REGION Network 21
   RUNG wire#powerrail
      { S7_Templates := "SrcType := String" } EQ_Contact(in1 := #String2, in2 := '6')
      Move(in := 125, out1 => #Decimal2_Out)
   END_RUNG
   // the same network as SCL:
   IF #String2 = '6' THEN #Decimal2_Out := 125; END_IF;
END_REGION

REGION Network 22
   RUNG wire#powerrail
      { S7_Templates := "SrcType := String" } EQ_Contact(in1 := #String2, in2 := '7')
      Move(in := 7, out1 => #Decimal2_Out)
   END_RUNG
   // the same network as SCL:
   IF #String2 = '7' THEN #Decimal2_Out := 7; END_IF;
END_REGION

REGION Network 23
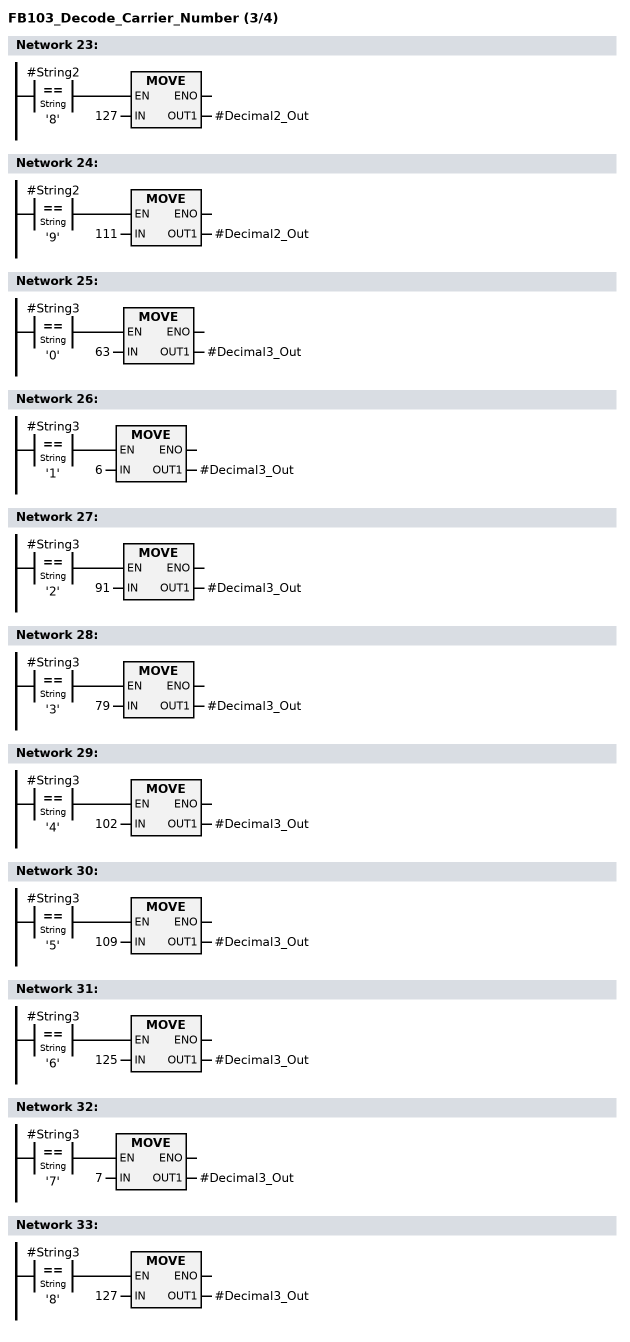
   RUNG wire#powerrail
      { S7_Templates := "SrcType := String" } EQ_Contact(in1 := #String2, in2 := '8')
      Move(in := 127, out1 => #Decimal2_Out)
   END_RUNG
   // the same network as SCL:
   IF #String2 = '8' THEN #Decimal2_Out := 127; END_IF;
END_REGION

REGION Network 24
   RUNG wire#powerrail
      { S7_Templates := "SrcType := String" } EQ_Contact(in1 := #String2, in2 := '9')
      Move(in := 111, out1 => #Decimal2_Out)
   END_RUNG
   // the same network as SCL:
   IF #String2 = '9' THEN #Decimal2_Out := 111; END_IF;
END_REGION

REGION Network 25
   RUNG wire#powerrail
      { S7_Templates := "SrcType := String" } EQ_Contact(in1 := #String3, in2 := '0')
      Move(in := 63, out1 => #Decimal3_Out)
   END_RUNG
   // the same network as SCL:
   IF #String3 = '0' THEN #Decimal3_Out := 63; END_IF;
END_REGION

REGION Network 26
   RUNG wire#powerrail
      { S7_Templates := "SrcType := String" } EQ_Contact(in1 := #String3, in2 := '1')
      Move(in := 6, out1 => #Decimal3_Out)
   END_RUNG
   // the same network as SCL:
   IF #String3 = '1' THEN #Decimal3_Out := 6; END_IF;
END_REGION

REGION Network 27
   RUNG wire#powerrail
      { S7_Templates := "SrcType := String" } EQ_Contact(in1 := #String3, in2 := '2')
      Move(in := 91, out1 => #Decimal3_Out)
   END_RUNG
   // the same network as SCL:
   IF #String3 = '2' THEN #Decimal3_Out := 91; END_IF;
END_REGION

REGION Network 28
   RUNG wire#powerrail
      { S7_Templates := "SrcType := String" } EQ_Contact(in1 := #String3, in2 := '3')
      Move(in := 79, out1 => #Decimal3_Out)
   END_RUNG
   // the same network as SCL:
   IF #String3 = '3' THEN #Decimal3_Out := 79; END_IF;
END_REGION

REGION Network 29
   RUNG wire#powerrail
      { S7_Templates := "SrcType := String" } EQ_Contact(in1 := #String3, in2 := '4')
      Move(in := 102, out1 => #Decimal3_Out)
   END_RUNG
   // the same network as SCL:
   IF #String3 = '4' THEN #Decimal3_Out := 102; END_IF;
END_REGION

REGION Network 30
   RUNG wire#powerrail
      { S7_Templates := "SrcType := String" } EQ_Contact(in1 := #String3, in2 := '5')
      Move(in := 109, out1 => #Decimal3_Out)
   END_RUNG
   // the same network as SCL:
   IF #String3 = '5' THEN #Decimal3_Out := 109; END_IF;
END_REGION

REGION Network 31
   RUNG wire#powerrail
      { S7_Templates := "SrcType := String" } EQ_Contact(in1 := #String3, in2 := '6')
      Move(in := 125, out1 => #Decimal3_Out)
   END_RUNG
   // the same network as SCL:
   IF #String3 = '6' THEN #Decimal3_Out := 125; END_IF;
END_REGION

REGION Network 32
   RUNG wire#powerrail
      { S7_Templates := "SrcType := String" } EQ_Contact(in1 := #String3, in2 := '7')
      Move(in := 7, out1 => #Decimal3_Out)
   END_RUNG
   // the same network as SCL:
   IF #String3 = '7' THEN #Decimal3_Out := 7; END_IF;
END_REGION

REGION Network 33
   RUNG wire#powerrail
      { S7_Templates := "SrcType := String" } EQ_Contact(in1 := #String3, in2 := '8')
      Move(in := 127, out1 => #Decimal3_Out)
   END_RUNG
   // the same network as SCL:
   IF #String3 = '8' THEN #Decimal3_Out := 127; END_IF;
END_REGION

REGION Network 34
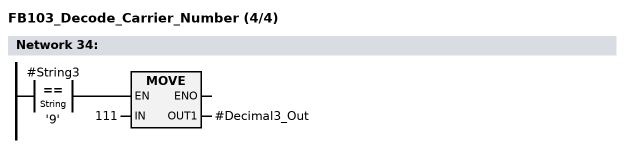
   RUNG wire#powerrail
      { S7_Templates := "SrcType := String" } EQ_Contact(in1 := #String3, in2 := '9')
      Move(in := 111, out1 => #Decimal3_Out)
   END_RUNG
   // the same network as SCL:
   IF #String3 = '9' THEN #Decimal3_Out := 111; END_IF;
END_REGION
END_FUNCTION_BLOCK

FUNCTION_BLOCK "FB104_CarrierBreakerStatus"   // FB104, LAD
{ S7_Optimized_Access := 'TRUE' }
AUTHOR : Siemens
VERSION : 1.0
// © 2018 Siemens AG 
// SIMOVE Carrier Control
   VAR
      instSystemBreakerStatus : "FB1001_EMS_BreakerStatus";
      instSystemDiagProfinet : "FB1003_LSimoveC_DiagProfinet";
      statCommunication : Bool;
      LSimoveC_DiagBreaker_Instance : "FB1001_EMS_BreakerStatus";
      LSimoveC_BreakerStatus_Instance : "FB1001_EMS_BreakerStatus";
   END_VAR
   VAR_TEMP
      tempBool_Tcc_2018_NotUsed : Bool;
   END_VAR
   VAR CONSTANT
      TCC2018_NotUsed : Bool;
   END_VAR
   VAR_TEMP   // added for the SCL form of the ladder/FBD networks
      _w1 : Bool;
   END_VAR
BEGIN

REGION Network 1: 10 System Monitoring Fuse
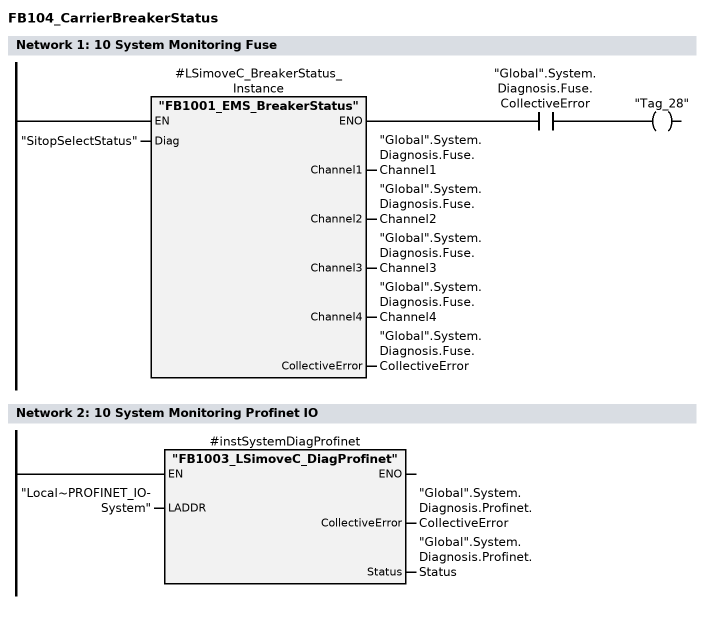
   RUNG wire#powerrail
      #LSimoveC_BreakerStatus_Instance(Diag := "SitopSelectStatus", Channel1 => "Global".System.Diagnosis.Fuse.Channel1, Channel2 => "Global".System.Diagnosis.Fuse.Channel2, Channel3 => "Global".System.Diagnosis.Fuse.Channel3, Channel4 => "Global".System.Diagnosis.Fuse.Channel4, CollectiveError => "Global".System.Diagnosis.Fuse.CollectiveError)
      Contact( "Global".System.Diagnosis.Fuse.CollectiveError )
      Coil( "Tag_28" )
   END_RUNG
   // the same network as SCL:
   #LSimoveC_BreakerStatus_Instance(Diag := "SitopSelectStatus",   // "FB1001_EMS_BreakerStatus"
                           Channel1 => "Global".System.Diagnosis.Fuse.Channel1,
                           Channel2 => "Global".System.Diagnosis.Fuse.Channel2,
                           Channel3 => "Global".System.Diagnosis.Fuse.Channel3,
                           Channel4 => "Global".System.Diagnosis.Fuse.Channel4,
                           CollectiveError => "Global".System.Diagnosis.Fuse.CollectiveError,
                           ENO => #_w1);
   "Tag_28" := #_w1 AND "Global".System.Diagnosis.Fuse.CollectiveError;
END_REGION

REGION Network 2: 10 System Monitoring Profinet IO
   RUNG wire#powerrail
      #instSystemDiagProfinet(LADDR := "Local~PROFINET_IO-System", CollectiveError => "Global".System.Diagnosis.Profinet.CollectiveError, Status => "Global".System.Diagnosis.Profinet.Status)
   END_RUNG
   // the same network as SCL:
   #instSystemDiagProfinet(LADDR := "Local~PROFINET_IO-System",   // "FB1003_LSimoveC_DiagProfinet"
                           CollectiveError => "Global".System.Diagnosis.Profinet.CollectiveError,
                           Status => "Global".System.Diagnosis.Profinet.Status);
END_REGION

REGION Network 3: 15 Navigation Transponder Antenna Left
END_REGION

REGION Network 4: 15 Navigation Transponder Antenna Right
END_REGION

REGION Network 5: 15 Navigation Identification Point
END_REGION
END_FUNCTION_BLOCK

FUNCTION_BLOCK "FB105_G120D_CarrierDrive"   // FB105, LAD
TITLE = Funkionblock for controlling a G120D
{ S7_Optimized_Access := 'FALSE' }
VERSION : 0.1
// -  ALLGEMEIN
//  - EINGÄNGE PEW
//  - STEUERWORT / CONTROLWORD
//  - ZUSTANDSWORT / STATUSWORD
//  - AUSGÄNGE PAW
//  - STÖRUNGEN
//  - ENDE
// 
// ________________________________________________________________________________
// 
// Groiß Andreas
// Siemens AG Österreich 
// Linz Kraußstraße 1-7 
// RC-AT I-IA AS-FA-SA-AE2
// 29.05.2013
// - GENERALLY
//  - INPUTS PEW
//  - STEUERWORT / CONTROLWORD
//  - ZUSTANDSWORT / STATUSWORD
//  - OUTPUTS PAW
//  - FAULTS
//  - END
// 
// ________________________________________________________________________________
// 
// Groiß Andreas
// Siemens AG Österreich 
// Linz Kraußstraße 1-7 
// I IA AS SO AP2 Surface Technology & Assembly
// 29.05.2013
   VAR_INPUT
      iPEW_ZSW1 : Word;   // IN: G120 D Zustandswort 1 / Stausword 1 PEW
      iPEW_SPEED : Word;   // IN: G120 D Aktual-Drehzahl / Actual-Speed of rotation PEW
      iPEW_INPUTS : Word;   // IN: G120 D digitale Eingänge / digital Inputs PEW
      iPEW_ERROR : Word;   // IN: G120 D Störcode / Errorcode PEW
      iEN_ERROR : Bool;   // IN: Freigabe Störmeldungen / IN: Enable Errormessages
      iON : Bool;   // IN: STW1_Bit_0 Steuerung Ein / IN: STW1_Bit_0 Control ON
      iPOWER_ON : Bool;   // IN: Kraftschalter ist EIN / IN: Power is switched on
      iENABLE : Bool;   // IN: Freigabe / IN: Enable
      iREVERSE : Bool;   // IN: STW1_Bit_11
      iBREAK : Bool;   // IN: Löse Bremse / IN: Release Break
      iDDS : Bool;   // IN: FU Datenset (0 = DDS0 / 1 = DDS1)
      iDO0 : Bool;   // IN: 1=Digitaler Ausgang aktiv/ 0=Digitaler Ausgang nicht aktiv
      iDO1 : Bool;   // IN: 1=Digitaler Ausgang aktiv/ 0=Digitaler Ausgang nicht aktiv
      iER_RESET : Bool;   // IN: Störung quittieren / IN: Error Reset
      iSET_SPEED : DInt;   // IN: Sollgeschwindigkeit in mm/min / IN: Setpoint Speed in mm/min
      iFACTOR : Real;   // IN: Übersetzungsfaktor m/min in Hz für G120D / IN: Conversion factor m/min in Hz for G120D
      iFACTOR_REV : Real;   // IN: Übersetzungsfaktor m/min in Hz für G120D reverse / IN: Conversion factor m/min in Hz for G120D reverse
      itON : Time;   // IN: TON ON
   END_VAR
   VAR_OUTPUT
      oPAW_STW1 : Word;   // OUT: G120 D Steuerwort 1 / Controlword 1 PAW
      oPAW_SPEED : Word;   // OUT: G120 D Soll-Drehzahl / Setpoint-Speed of rotation PAW
      oCUR_SPEED : DInt;   // OUT: G120 D Current speed in mm/min
      oZSW1 : "UDT_G120D_ZSW1_STATUS";   // OUT: G120 D Zustandswort 1 / Stausword 1
      oSTW1 : "UDT_G120D_STW1_CONTROL";   // OUT: G120 D Steuerwort 1 / Controlword 1
      oINPUTS : Struct   // OUT: G120 D Eingänge / Inputs
         E_1_0 : Bool;   // G120 D Eingänge / Inputs 1.0
         E_1_1 : Bool;   // G120 D Eingänge / Inputs 1.1
         E_1_2 : Bool;   // G120 D Eingänge / Inputs 1.2
         E_1_3 : Bool;   // G120 D Eingänge / Inputs 1.3
         E_1_4 : Bool;   // G120 D Eingänge / Inputs 1.4
         E_1_5 : Bool;   // G120 D Eingänge / Inputs 1.5
         E_1_6 : Bool;   // G120 D Eingänge / Inputs 1.6
         E_1_7 : Bool;   // G120 D Eingänge / Inputs 1.7
         E_0_0 : Bool;   // G120 D Eingänge / Inputs 0.0
         E_0_1 : Bool;   // G120 D Eingänge / Inputs 0.1
         E_0_2 : Bool;   // G120 D Eingänge / Inputs 0.2
         E_0_3 : Bool;   // G120 D Eingänge / Inputs 0.3
         E_0_4 : Bool;   // G120 D Eingänge / Inputs 0.4
         E_0_5 : Bool;   // G120 D Eingänge / Inputs 0.5
         E_0_6 : Bool;   // G120 D Eingänge / Inputs 0.6
         E_0_7 : Bool;   // G120 D Eingänge / Inputs 0.7
      END_STRUCT;
      oER_FC : Bool;   // OUT: Störung FU allgemein / OUT: Error / ZSW1_Bit_3
      oER_SUM : Bool;   // OUT: Sammelstörung / OUT: Error Summary
   END_VAR
   VAR_IN_OUT
      ioERRORS : Struct   // INOUT: G120D Störungen / INOUT: G120D Faults
         ER000 : Bool;   // INOUT: Störung XXX / INOUT: Error XXX
         ER001 : Bool;   // INOUT: Störung XXX / INOUT: Error XXX
         ER002 : Bool;   // INOUT: Störung XXX / INOUT: Error XXX
         ER003 : Bool;   // INOUT: Störung XXX / INOUT: Error XXX
         ER004 : Bool;   // INOUT: Störung XXX / INOUT: Error XXX
         ER005 : Bool;   // INOUT: Störung XXX / INOUT: Error XXX
         ER006 : Bool;   // INOUT: Störung XXX / INOUT: Error XXX
         ER007 : Bool;   // INOUT: Störung XXX / INOUT: Error XXX
         ER008 : Bool;   // INOUT: Störung XXX / INOUT: Error XXX
         ER009 : Bool;   // INOUT: Störung XXX / INOUT: Error XXX
         ER010 : Bool;   // INOUT: Störung XXX / INOUT: Error XXX
         ER011 : Bool;   // INOUT: Störung XXX / INOUT: Error XXX
         ER012 : Bool;   // INOUT: Störung XXX / INOUT: Error XXX
         ER013 : Bool;   // INOUT: Störung XXX / INOUT: Error XXX
         ER014 : Bool;   // INOUT: Störung XXX / INOUT: Error XXX
         ER015 : Bool;   // INOUT: Störung XXX / INOUT: Error XXX
      END_STRUCT;
      ioERROR_PAR : Struct
         ER000 : Int;   // INOUT: Störnummer XXX / INOUT: Error Number XXX
         ER001 : Int;   // INOUT: Störnummer XXX / INOUT: Error Number XXX
         ER002 : Int;   // INOUT: Störnummer XXX / INOUT: Error Number XXX
         ER003 : Int;   // INOUT: Störnummer XXX / INOUT: Error Number XXX
         ER004 : Int;   // INOUT: Störnummer XXX / INOUT: Error Number XXX
         ER005 : Int;   // INOUT: Störnummer XXX / INOUT: Error Number XXX
         ER006 : Int;   // INOUT: Störnummer XXX / INOUT: Error Number XXX
         ER007 : Int;   // INOUT: Störnummer XXX / INOUT: Error Number XXX
         ER008 : Int;   // INOUT: Störnummer XXX / INOUT: Error Number XXX
         ER009 : Int;   // INOUT: Störnummer XXX / INOUT: Error Number XXX
         ER010 : Int;   // INOUT: Störnummer XXX / INOUT: Error Number XXX
         ER011 : Int;   // INOUT: Störnummer XXX / INOUT: Error Number XXX
         ER012 : Int;   // INOUT: Störnummer XXX / INOUT: Error Number XXX
         ER013 : Int;   // INOUT: Störnummer XXX / INOUT: Error Number XXX
         ER014 : Int;   // INOUT: Störnummer XXX / INOUT: Error Number XXX
         ER015 : Int;   // INOUT: Störnummer XXX / INOUT: Error Number XXX
      END_STRUCT;
   END_VAR
   VAR
      STAT_MI_EN_Faults : TON_TIME;   // STAT: TON Freigabe Störungen / STAT: TON enable Faults
      STAT_MI_On : TON_TIME;   // STAT: TON EIN / STAT: TON On
      STAT_MI_TP_Reset : IEC_TIMER;   // STAT: TP Rücksetzen
      STAT_MI_TON_Reset : IEC_TIMER;   // STAT: TON Rücksetzen
      STAT_MI_TOF_On : IEC_TIMER;   // STAT: TOF EIN
      STAT_oER_FC : Bool;   // STAT: Störung FU allgemein / OUT: Error / ZSW1_Bit_3
   END_VAR
   VAR_TEMP
      Temp_SEND : Struct   // TEMP: sende LW 0 !!! nicht verschieben !!! / TEMP: send LW 0 !!! don`t move !!!
         STW1 : Struct   // TEMP: G120 D Steuerwort 1 / Controlword 1 !!! LW0 don`t move !!!
            Bit_08_JOG_R : Bool;   // 1=jogging on right-hand side ON/ 0= OFF
            Bit_09_JOG_L : Bool;   // 1=jogging on left-hand side ON/ 0= OFF
            Bit_10_CONTR_PLC : Bool;   // 1=control by PLC required/ 0=no control by PLC required
            Bit_11_REVERSE : Bool;   // 1=inversion of setpoint/ 0=no inversion of setpoint
            Bit_12_BREAK : Bool;   // 1= Release Break
            Bit_13_DDS : Bool;   // 1=DDS1 FU Dataset / 0=DDS0 FU Dataset / 1=Motor potentiometer up ON/ 0=OFF
            Bit_14_DO0 : Bool;   // 1=Digital Output activ/ 0=Digital Output not activ / 1=Motor potentiometer down ON/ 0=OFF
            Bit_15_DO1 : Bool;   // 1=Digital Output activ/ 0=Digital Output not activ / 1=local control (BOP/AOP) active/ 0=remote control active
            Bit_00_ON : Bool;   // 1=ON/ 0=OFF2 / 1=ON/ 0=OFF1
            Bit_01_AUS2_INH : Bool;   // 1=operation condition/ 0=AUS2 - pulse inhibitor, voltage off at once
            Bit_02_AUS3_STOP : Bool;   // 1=operation condition / 0=AUS3 - fast stop
            Bit_03_EN : Bool;   // 1=enable operation/ 0=disable operation
            Bit_04_EN_RAMP : Bool;   // 1=operation condition / 0=disable ramp function generator
            Bit_05_START_RAMP : Bool;   // 1=enable ramp function generator / 0=stoppen RFG
            Bit_06_SETPOINT : Bool;   // 1=enable setpoint/ 0=disable setpoint
            Bit_07_RESET : Bool;   // 1=Reset fault / 0= irrelevant
         END_STRUCT;
         SPEED : Word;   // TEMP: G120 D Soll-Drehzahl / Setpoint-Speed of rotation !!! LW2 don`t move !!!
         SPARE : Array[4..9] of Byte;   // TEMP: Spare !!! LW4 don`t move !!!
      END_STRUCT;
      Temp_REC : Struct   // TEMP: empfange LW 10 !!! nicht verschieben !!! / TEMP: receive LW 10 !!! don`t move !!!
         ZSW1 : Struct   // TEMP: G120 D Zustandswort 1 / Stausword 1 !!! LW10 don`t move !!!
            Bit_08_NO_DEVIATION : Bool;   // 1=no deviation current-setpoint / 0=deviation
            Bit_09_CONTR_PLC : Bool;   // 1=control by PLC required/ 0=no control by PLC required
            Bit_10_F_MAX : Bool;   // 1=fmax reached/ 0= below fmax
            Bit_11_NO_WARN : Bool;   // 1=no warning/ 0=warning:Motor at limit of current
            Bit_12_NO_BREAK : Bool;   // 1= / 0=Haltebremse
            Bit_13_NO_OVERL : Bool;   // 1= / 0=Motorüberlast
            Bit_14_CW_CCW : Bool;   // 1=Rechtslauf/ 0=Linkslauf
            Bit_15_OVERL : Bool;   // 1= /0= Konverter overload
            Bit_00_READY_RUN : Bool;   // 1=ready to run/ 0= not ready to run
            Bit_01_READY_ON : Bool;   // 1=ready to switch on/ 0= not ready to switch on
            Bit_02_ENABLE : Bool;   // 1=operation enabled / 0=operation disabled
            Bit_03_FAULT : Bool;   // 1=fault / 0=no fault
            Bit_04_AUS2 : Bool;   // 1=no AUS2 / 0=AUS2 command is present
            Bit_05_AUS3 : Bool;   // 1=no AUS3 / 0=AUS3 command is present
            Bit_06_LOCK_OUT : Bool;   // 1=closing lock-out / 0=no closing lock-out
            Bit_07_WARN : Bool;   // 1=Warning / 0= no warning
         END_STRUCT;
         SPEED : Int;   // TEMP: G120 D Aktuel-Drehzahl / Actual-Speed of rotation !!! LW12 don`t move !!!
         INPUTS : Struct   // TEMP: G120 D Eingänge / Inputs !!! LW14 don`t move !!!
            I_XX1_0 : Bool;   // G120 D Eingänge / Inputs XX1.0
            I_XX1_1 : Bool;   // G120 D Eingänge / Inputs XX1.1
            I_XX1_2 : Bool;   // G120 D Eingänge / Inputs XX1.2
            I_XX1_3 : Bool;   // G120 D Eingänge / Inputs XX1.3
            I_XX1_4 : Bool;   // G120 D Eingänge / Inputs XX1.4
            I_XX1_5 : Bool;   // G120 D Eingänge / Inputs XX1.5
            I_XX1_6 : Bool;   // G120 D Eingänge / Inputs XX1.6
            I_XX1_7 : Bool;   // G120 D Eingänge / Inputs XX1.7
            I_XX0_0 : Bool;   // G120 D Eingänge / Inputs XX0.0
            I_XX0_1 : Bool;   // G120 D Eingänge / Inputs XX0.1
            I_XX0_2 : Bool;   // G120 D Eingänge / Inputs XX0.2
            I_XX0_3 : Bool;   // G120 D Eingänge / Inputs XX0.3
            I_XX0_4 : Bool;   // G120 D Eingänge / Inputs XX0.4
            I_XX0_5 : Bool;   // G120 D Eingänge / Inputs XX0.5
            I_XX0_6 : Bool;   // G120 D Eingänge / Inputs XX0.6
            I_XX0_7 : Bool;   // G120 D Eingänge / Inputs XX0.7
         END_STRUCT;
         ERROR : Int;   // TEMP: G120 D Störcode / Errorcode !!! LW16 don`t move !!! / TEMP: G120 D Störcode / Faultcode !!! LW16 don`t move !!!
         SPARE : Array[18..19] of Byte;   // TEMP: Spare !!! LW4 don`t move !!!
      END_STRUCT;
      Temp_AR1 : DWord;   // TEMP: AR1
      Temp_AR2 : DWord;   // TEMP: AR2
      Temp_Real : Real;   // TEMP: Temprärer Speicher / TEMP: Temporary memory
      Temp_RetVal : Int;   // TEMP: RetVal
      Temp_Factor : Real;   // TEMP: Faktor / TEMP: Factor
      Temp_Int_0 : Int;   // TEMP: Null
      Temp_Null : Bool;   // TEMP: feste Null
      Temp_Eins : Bool;   // TEMP: feste Eins
      Temp_ON : Bool;   // TEMP: ON
      Temp_EN_Faults : Bool;   // TEMP: Freigabe Fehler / TEMP: Enable Faults
   END_VAR
   VAR_TEMP   // added for the SCL form of the ladder/FBD networks
      _w1 : Bool;
   END_VAR
BEGIN

REGION Network 1: ALLGEMEIN / GENERALLY
   // ################################## ALLGEMEIN ########################## / ################################## GENERALLY ##################################
END_REGION

REGION Network 2: TEMP: feste Eins / Null
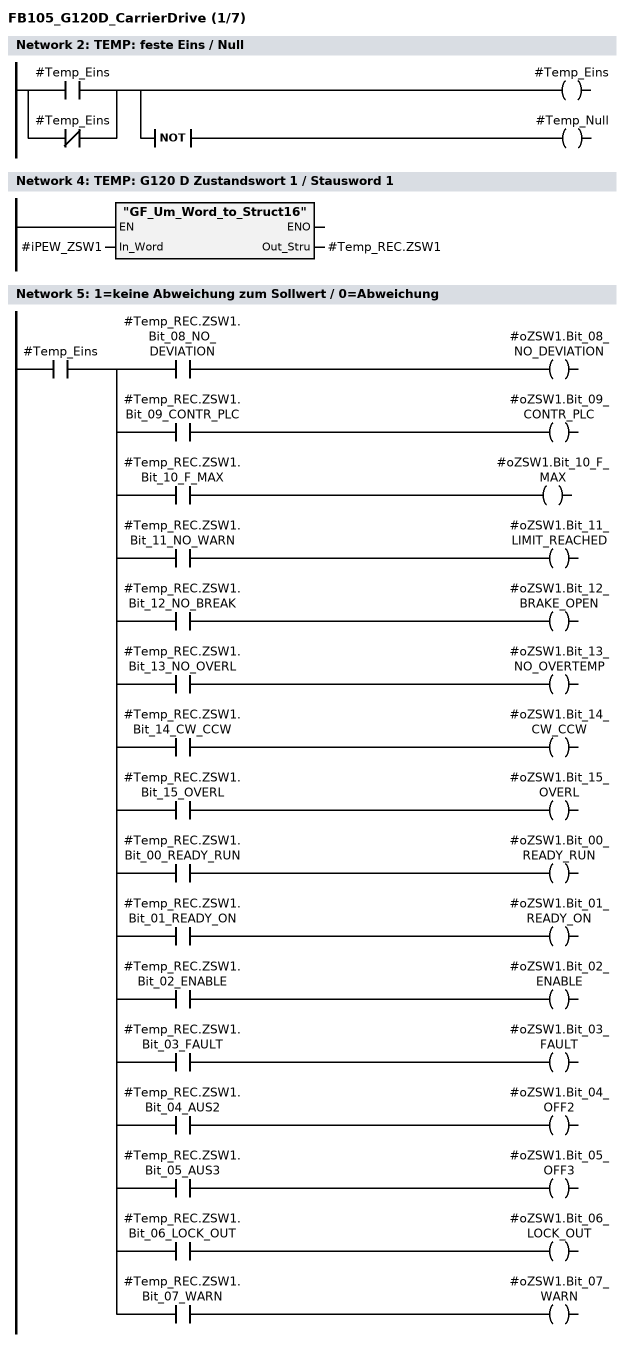
   RUNG wire#powerrail
      Contact( #Temp_Eins )
      wire#w1
      Coil( #Temp_Eins )
   END_RUNG
   RUNG wire#powerrail
      I_Contact( #Temp_Eins )
   END_RUNG wire#w1
   RUNG wire#w1
      Not()
      Coil( #Temp_Null )
   END_RUNG
   // the same network as SCL:
   #Temp_Eins := #Temp_Eins OR NOT #Temp_Eins;
   #Temp_Null := NOT #Temp_Eins;
END_REGION

REGION Network 3: EINGÄNGE PEW / INPUTS PEW
   // ##################################### PEW ######################################
END_REGION

REGION Network 4: TEMP: G120 D Zustandswort 1 / Stausword 1
   RUNG wire#powerrail
      "GF_Um_Word_to_Struct16"(In_Word := #iPEW_ZSW1, Out_Stru => #Temp_REC.ZSW1)
   END_RUNG
   // the same network as SCL:
   "GF_Um_Word_to_Struct16"(In_Word := #iPEW_ZSW1, Out_Stru => #Temp_REC.ZSW1);
END_REGION

REGION Network 5: 1=keine Abweichung zum Sollwert / 0=Abweichung
   RUNG wire#powerrail
      Contact( #Temp_Eins )
      wire#w1
      Contact( #Temp_REC.ZSW1.Bit_08_NO_DEVIATION )
      Coil( #oZSW1.Bit_08_NO_DEVIATION )
   END_RUNG
   RUNG wire#w1
      Contact( #Temp_REC.ZSW1.Bit_09_CONTR_PLC )
      Coil( #oZSW1.Bit_09_CONTR_PLC )
   END_RUNG
   RUNG wire#w1
      Contact( #Temp_REC.ZSW1.Bit_10_F_MAX )
      Coil( #oZSW1.Bit_10_F_MAX )
   END_RUNG
   RUNG wire#w1
      Contact( #Temp_REC.ZSW1.Bit_11_NO_WARN )
      Coil( #oZSW1.Bit_11_LIMIT_REACHED )
   END_RUNG
   RUNG wire#w1
      Contact( #Temp_REC.ZSW1.Bit_12_NO_BREAK )
      Coil( #oZSW1.Bit_12_BRAKE_OPEN )
   END_RUNG
   RUNG wire#w1
      Contact( #Temp_REC.ZSW1.Bit_13_NO_OVERL )
      Coil( #oZSW1.Bit_13_NO_OVERTEMP )
   END_RUNG
   RUNG wire#w1
      Contact( #Temp_REC.ZSW1.Bit_14_CW_CCW )
      Coil( #oZSW1.Bit_14_CW_CCW )
   END_RUNG
   RUNG wire#w1
      Contact( #Temp_REC.ZSW1.Bit_15_OVERL )
      Coil( #oZSW1.Bit_15_OVERL )
   END_RUNG
   RUNG wire#w1
      Contact( #Temp_REC.ZSW1.Bit_00_READY_RUN )
      Coil( #oZSW1.Bit_00_READY_RUN )
   END_RUNG
   RUNG wire#w1
      Contact( #Temp_REC.ZSW1.Bit_01_READY_ON )
      Coil( #oZSW1.Bit_01_READY_ON )
   END_RUNG
   RUNG wire#w1
      Contact( #Temp_REC.ZSW1.Bit_02_ENABLE )
      Coil( #oZSW1.Bit_02_ENABLE )
   END_RUNG
   RUNG wire#w1
      Contact( #Temp_REC.ZSW1.Bit_03_FAULT )
      Coil( #oZSW1.Bit_03_FAULT )
   END_RUNG
   RUNG wire#w1
      Contact( #Temp_REC.ZSW1.Bit_04_AUS2 )
      Coil( #oZSW1.Bit_04_OFF2 )
   END_RUNG
   RUNG wire#w1
      Contact( #Temp_REC.ZSW1.Bit_05_AUS3 )
      Coil( #oZSW1.Bit_05_OFF3 )
   END_RUNG
   RUNG wire#w1
      Contact( #Temp_REC.ZSW1.Bit_06_LOCK_OUT )
      Coil( #oZSW1.Bit_06_LOCK_OUT )
   END_RUNG
   RUNG wire#w1
      Contact( #Temp_REC.ZSW1.Bit_07_WARN )
      Coil( #oZSW1.Bit_07_WARN )
   END_RUNG
   // the same network as SCL:
   #oZSW1.Bit_08_NO_DEVIATION := #Temp_Eins AND #Temp_REC.ZSW1.Bit_08_NO_DEVIATION;
   #oZSW1.Bit_09_CONTR_PLC := #Temp_Eins AND #Temp_REC.ZSW1.Bit_09_CONTR_PLC;
   #oZSW1.Bit_10_F_MAX := #Temp_Eins AND #Temp_REC.ZSW1.Bit_10_F_MAX;
   #oZSW1.Bit_11_LIMIT_REACHED := #Temp_Eins AND #Temp_REC.ZSW1.Bit_11_NO_WARN;
   #oZSW1.Bit_12_BRAKE_OPEN := #Temp_Eins AND #Temp_REC.ZSW1.Bit_12_NO_BREAK;
   #oZSW1.Bit_13_NO_OVERTEMP := #Temp_Eins AND #Temp_REC.ZSW1.Bit_13_NO_OVERL;
   #oZSW1.Bit_14_CW_CCW := #Temp_Eins AND #Temp_REC.ZSW1.Bit_14_CW_CCW;
   #oZSW1.Bit_15_OVERL := #Temp_Eins AND #Temp_REC.ZSW1.Bit_15_OVERL;
   #oZSW1.Bit_00_READY_RUN := #Temp_Eins AND #Temp_REC.ZSW1.Bit_00_READY_RUN;
   #oZSW1.Bit_01_READY_ON := #Temp_Eins AND #Temp_REC.ZSW1.Bit_01_READY_ON;
   #oZSW1.Bit_02_ENABLE := #Temp_Eins AND #Temp_REC.ZSW1.Bit_02_ENABLE;
   #oZSW1.Bit_03_FAULT := #Temp_Eins AND #Temp_REC.ZSW1.Bit_03_FAULT;
   #oZSW1.Bit_04_OFF2 := #Temp_Eins AND #Temp_REC.ZSW1.Bit_04_AUS2;
   #oZSW1.Bit_05_OFF3 := #Temp_Eins AND #Temp_REC.ZSW1.Bit_05_AUS3;
   #oZSW1.Bit_06_LOCK_OUT := #Temp_Eins AND #Temp_REC.ZSW1.Bit_06_LOCK_OUT;
   #oZSW1.Bit_07_WARN := #Temp_Eins AND #Temp_REC.ZSW1.Bit_07_WARN;
END_REGION

REGION Network 6: TEMP: G120 D Eingänge / Inputs
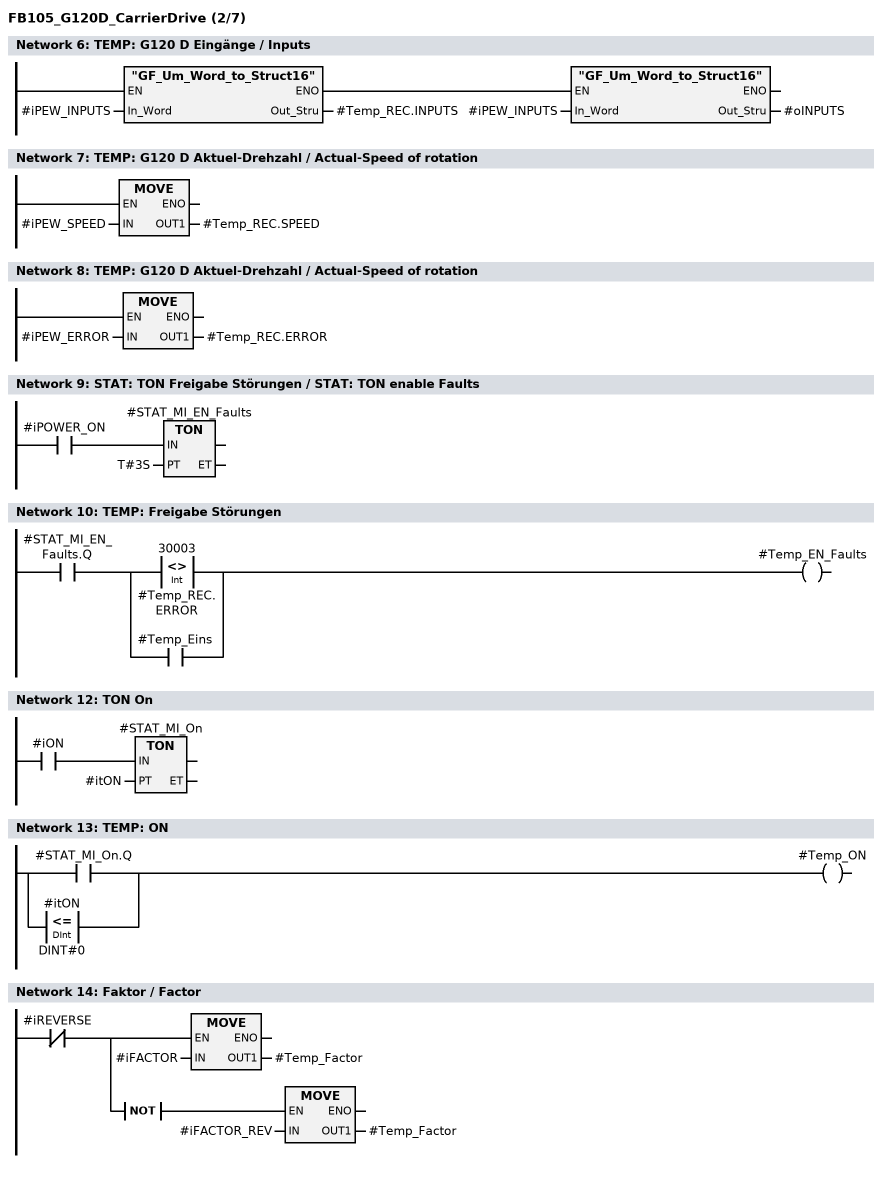
   RUNG wire#powerrail
      "GF_Um_Word_to_Struct16"(In_Word := #iPEW_INPUTS, Out_Stru => #Temp_REC.INPUTS)
      "GF_Um_Word_to_Struct16"(In_Word := #iPEW_INPUTS, Out_Stru => #oINPUTS)
   END_RUNG
   // the same network as SCL:
   "GF_Um_Word_to_Struct16"(In_Word := #iPEW_INPUTS, Out_Stru => #Temp_REC.INPUTS, ENO => #_w1);
   IF #_w1 THEN "GF_Um_Word_to_Struct16"(In_Word := #iPEW_INPUTS, Out_Stru => #oINPUTS); END_IF;
END_REGION

REGION Network 7: TEMP: G120 D Aktuel-Drehzahl / Actual-Speed of rotation
   RUNG wire#powerrail
      Move(in := #iPEW_SPEED, out1 => #Temp_REC.SPEED)
   END_RUNG
   // the same network as SCL:
   #Temp_REC.SPEED := #iPEW_SPEED;
END_REGION

REGION Network 8: TEMP: G120 D Aktuel-Drehzahl / Actual-Speed of rotation
   RUNG wire#powerrail
      Move(in := #iPEW_ERROR, out1 => #Temp_REC.ERROR)
   END_RUNG
   // the same network as SCL:
   #Temp_REC.ERROR := #iPEW_ERROR;
END_REGION

REGION Network 9: STAT: TON Freigabe Störungen / STAT: TON enable Faults
   #STAT_MI_EN_Faults(IN := #iPOWER_ON, PT := T#3S);   // TON
END_REGION

REGION Network 10: TEMP: Freigabe Störungen
   RUNG wire#powerrail
      Contact( #STAT_MI_EN_Faults.Q )
      wire#w1
      { S7_Templates := "SrcType := Int" } NE_Contact(in1 := 30003, in2 := #Temp_REC.ERROR)
      wire#w2
      Coil( #Temp_EN_Faults )
   END_RUNG
   RUNG wire#w1
      Contact( #Temp_Eins )
   END_RUNG wire#w2
   // the same network as SCL:
   #Temp_EN_Faults := #STAT_MI_EN_Faults.Q AND ((30003 <> #Temp_REC.ERROR) OR #Temp_Eins);
END_REGION

REGION Network 11: STEUERWORT / CONTROLWORD
   // ##################################### STW #####################################
END_REGION

REGION Network 12: TON On
   #STAT_MI_On(IN := #iON, PT := #itON);   // TON
END_REGION

REGION Network 13: TEMP: ON
   RUNG wire#powerrail
      Contact( #STAT_MI_On.Q )
      wire#w1
      Coil( #Temp_ON )
   END_RUNG
   RUNG wire#powerrail
      { S7_Templates := "SrcType := DInt" } LE_Contact(in1 := #itON, in2 := DINT#0)
   END_RUNG wire#w1
   // the same network as SCL:
   #Temp_ON := #STAT_MI_On.Q OR (#itON <= DINT#0);
END_REGION

REGION Network 14: Faktor / Factor
   RUNG wire#powerrail
      I_Contact( #iREVERSE )
      wire#w1
      { S7_GenerateENO := "TRUE" } Move(in := #iFACTOR, out1 => #Temp_Factor)
   END_RUNG
   RUNG wire#w1
      Not()
      { S7_GenerateENO := "TRUE" } Move(in := #iFACTOR_REV, out1 => #Temp_Factor)
   END_RUNG
   // the same network as SCL:
   IF NOT #iREVERSE THEN #Temp_Factor := #iFACTOR; END_IF;
   IF NOT (NOT #iREVERSE) THEN #Temp_Factor := #iFACTOR_REV; END_IF;
END_REGION

REGION Network 15 (STL): Generiere Befehle und Sollwerte / Generate control commands and setpoint
         SET;  // Setzt VKE=1
         =     #Temp_SEND.STW1.Bit_01_AUS2_INH;
         =     #Temp_SEND.STW1.Bit_04_EN_RAMP;
         =     #Temp_SEND.STW1.Bit_05_START_RAMP;
         =     #Temp_SEND.STW1.Bit_06_SETPOINT;
         =     #Temp_SEND.STW1.Bit_10_CONTR_PLC;  // Führung AG gefordert !!

         CLR;  // Setzt VKE=0
         =     #Temp_SEND.STW1.Bit_08_JOG_R;
         =     #Temp_SEND.STW1.Bit_09_JOG_L;

         A     #Temp_ON;  // Abfrage der Bausteinschnittstelle
         A     #Temp_REC.ZSW1.Bit_00_READY_RUN;  // Antrieb bereit
         A     #iPOWER_ON;
         A     #iEN_ERROR;
         =     #Temp_SEND.STW1.Bit_00_ON;

         A     #STAT_MI_TOF_On.Q;
         O     #Temp_SEND.STW1.Bit_00_ON;
         =     #Temp_SEND.STW1.Bit_03_EN;

         A     #iENABLE;
         =     #Temp_SEND.STW1.Bit_02_AUS3_STOP;

         A     #iREVERSE;
         =     #Temp_SEND.STW1.Bit_11_REVERSE;

         A     #iBREAK;
         =     #Temp_SEND.STW1.Bit_12_BREAK;

         A     #iDDS;
         =     #Temp_SEND.STW1.Bit_13_DDS;  // Datensatzumschaltung

         A     #iDO0;
         =     #Temp_SEND.STW1.Bit_14_DO0;  // Ausgang DO0 z.B.: Ansteuerung Meldelampe

         A     #iDO1;
         =     #Temp_SEND.STW1.Bit_15_DO1;  // Ausgang DO1 z.B.: Ansteuerung Staubsauger

   //
   // PZD2 - Drehzahlsollwert
   // gültiger Drehzahlsollwert zwischen 0.00-130 % (% bezogen auf Bezugsdrehzhal in FU

         L     #iSET_SPEED;
         DTR;
         L     #Temp_Factor;
         *R;
         T     #Temp_Real;  // Frequenzsollwert [%]

         L     0.0;
         >R;  // Drehzahlsollwert <0%
         JC    N010;
         T     #Temp_Real;  // Frequenzsollwert [%]

   N010: L     #Temp_Real;  // Frequenzsollwert [%]
         L     130.0;
         <R;  // Drehzahlsollwert >130% ?
         JC    N011;
         T     #Temp_Real;  // Frequenzsollwert [%]

   N011: L     #Temp_Real;  // Frequenzsollwert [%]
         L     100.0;  // 2-Nachkommastellen retten
         *R;
         RND;  // Umwandeln 32Bit Realzahl in 32Bit Ganzzahl
         L     16384;  // 16384 = 4000HEX = 100%
         *D;
         L     10000;
         /D;
         T     #Temp_SEND.SPEED;  // Transfer in das Sendefach

         NOP   0;
END_REGION

REGION Network 16: Generiere Befehle Neustart
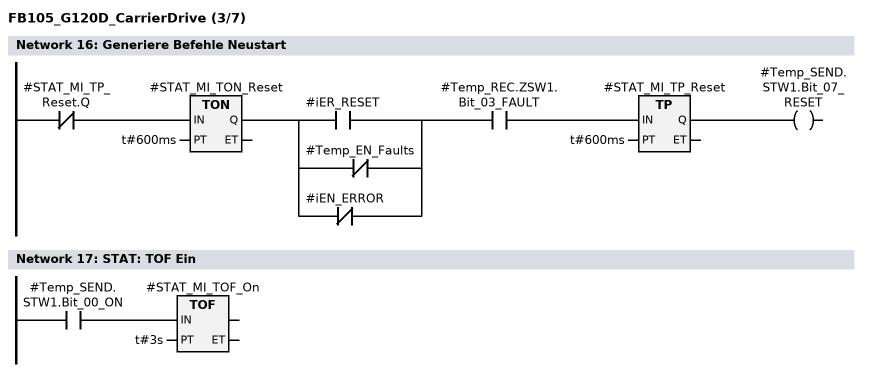
   #STAT_MI_TON_Reset.TON(IN := NOT #STAT_MI_TP_Reset.Q, PT := t#600ms);
   #STAT_MI_TP_Reset.TP(IN := #STAT_MI_TON_Reset.Q AND (#iER_RESET OR NOT #Temp_EN_Faults OR NOT #iEN_ERROR) AND #Temp_REC.ZSW1.Bit_03_FAULT,
                        PT := t#600ms);
   #Temp_SEND.STW1.Bit_07_RESET := #STAT_MI_TP_Reset.Q;
END_REGION

REGION Network 17: STAT: TOF Ein
   #STAT_MI_TOF_On.TOF(IN := #Temp_SEND.STW1.Bit_00_ON, PT := t#3s);
END_REGION

REGION Network 18: STW
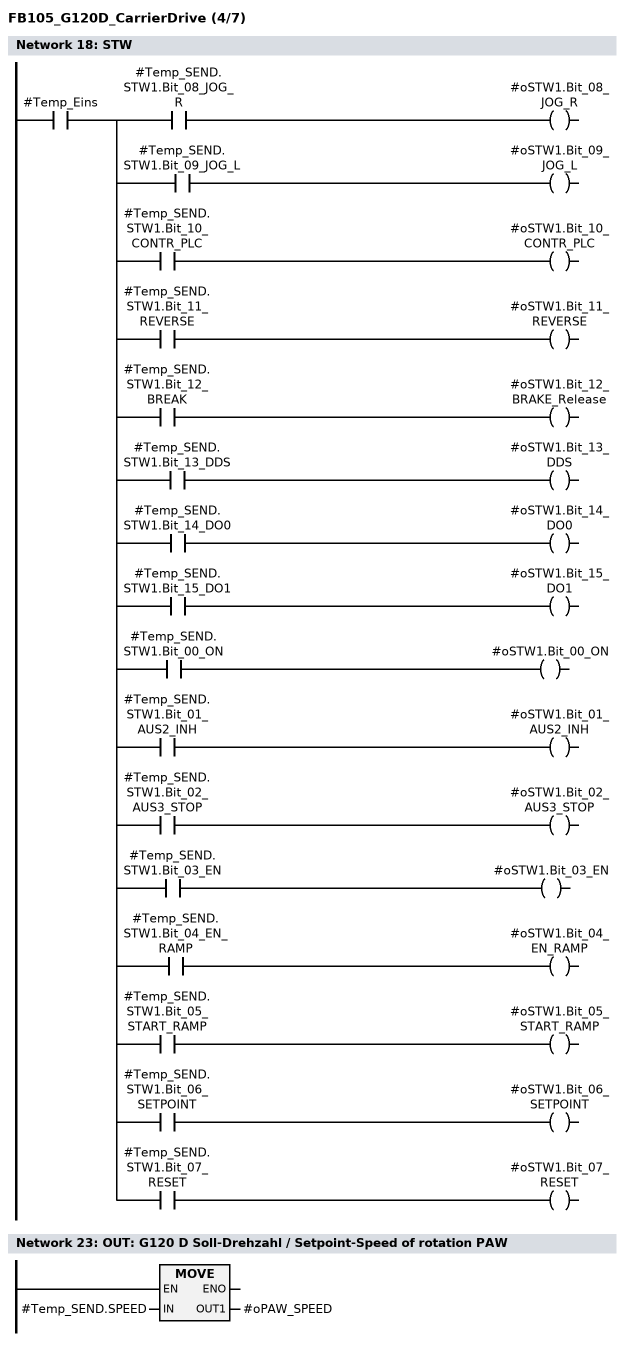
   RUNG wire#powerrail
      Contact( #Temp_Eins )
      wire#w1
      Contact( #Temp_SEND.STW1.Bit_08_JOG_R )
      Coil( #oSTW1.Bit_08_JOG_R )
   END_RUNG
   RUNG wire#w1
      Contact( #Temp_SEND.STW1.Bit_09_JOG_L )
      Coil( #oSTW1.Bit_09_JOG_L )
   END_RUNG
   RUNG wire#w1
      Contact( #Temp_SEND.STW1.Bit_10_CONTR_PLC )
      Coil( #oSTW1.Bit_10_CONTR_PLC )
   END_RUNG
   RUNG wire#w1
      Contact( #Temp_SEND.STW1.Bit_11_REVERSE )
      Coil( #oSTW1.Bit_11_REVERSE )
   END_RUNG
   RUNG wire#w1
      Contact( #Temp_SEND.STW1.Bit_12_BREAK )
      Coil( #oSTW1.Bit_12_BRAKE_Release )
   END_RUNG
   RUNG wire#w1
      Contact( #Temp_SEND.STW1.Bit_13_DDS )
      Coil( #oSTW1.Bit_13_DDS )
   END_RUNG
   RUNG wire#w1
      Contact( #Temp_SEND.STW1.Bit_14_DO0 )
      Coil( #oSTW1.Bit_14_DO0 )
   END_RUNG
   RUNG wire#w1
      Contact( #Temp_SEND.STW1.Bit_15_DO1 )
      Coil( #oSTW1.Bit_15_DO1 )
   END_RUNG
   RUNG wire#w1
      Contact( #Temp_SEND.STW1.Bit_00_ON )
      Coil( #oSTW1.Bit_00_ON )
   END_RUNG
   RUNG wire#w1
      Contact( #Temp_SEND.STW1.Bit_01_AUS2_INH )
      Coil( #oSTW1.Bit_01_AUS2_INH )
   END_RUNG
   RUNG wire#w1
      Contact( #Temp_SEND.STW1.Bit_02_AUS3_STOP )
      Coil( #oSTW1.Bit_02_AUS3_STOP )
   END_RUNG
   RUNG wire#w1
      Contact( #Temp_SEND.STW1.Bit_03_EN )
      Coil( #oSTW1.Bit_03_EN )
   END_RUNG
   RUNG wire#w1
      Contact( #Temp_SEND.STW1.Bit_04_EN_RAMP )
      Coil( #oSTW1.Bit_04_EN_RAMP )
   END_RUNG
   RUNG wire#w1
      Contact( #Temp_SEND.STW1.Bit_05_START_RAMP )
      Coil( #oSTW1.Bit_05_START_RAMP )
   END_RUNG
   RUNG wire#w1
      Contact( #Temp_SEND.STW1.Bit_06_SETPOINT )
      Coil( #oSTW1.Bit_06_SETPOINT )
   END_RUNG
   RUNG wire#w1
      Contact( #Temp_SEND.STW1.Bit_07_RESET )
      Coil( #oSTW1.Bit_07_RESET )
   END_RUNG
   // the same network as SCL:
   #oSTW1.Bit_08_JOG_R := #Temp_Eins AND #Temp_SEND.STW1.Bit_08_JOG_R;
   #oSTW1.Bit_09_JOG_L := #Temp_Eins AND #Temp_SEND.STW1.Bit_09_JOG_L;
   #oSTW1.Bit_10_CONTR_PLC := #Temp_Eins AND #Temp_SEND.STW1.Bit_10_CONTR_PLC;
   #oSTW1.Bit_11_REVERSE := #Temp_Eins AND #Temp_SEND.STW1.Bit_11_REVERSE;
   #oSTW1.Bit_12_BRAKE_Release := #Temp_Eins AND #Temp_SEND.STW1.Bit_12_BREAK;
   #oSTW1.Bit_13_DDS := #Temp_Eins AND #Temp_SEND.STW1.Bit_13_DDS;
   #oSTW1.Bit_14_DO0 := #Temp_Eins AND #Temp_SEND.STW1.Bit_14_DO0;
   #oSTW1.Bit_15_DO1 := #Temp_Eins AND #Temp_SEND.STW1.Bit_15_DO1;
   #oSTW1.Bit_00_ON := #Temp_Eins AND #Temp_SEND.STW1.Bit_00_ON;
   #oSTW1.Bit_01_AUS2_INH := #Temp_Eins AND #Temp_SEND.STW1.Bit_01_AUS2_INH;
   #oSTW1.Bit_02_AUS3_STOP := #Temp_Eins AND #Temp_SEND.STW1.Bit_02_AUS3_STOP;
   #oSTW1.Bit_03_EN := #Temp_Eins AND #Temp_SEND.STW1.Bit_03_EN;
   #oSTW1.Bit_04_EN_RAMP := #Temp_Eins AND #Temp_SEND.STW1.Bit_04_EN_RAMP;
   #oSTW1.Bit_05_START_RAMP := #Temp_Eins AND #Temp_SEND.STW1.Bit_05_START_RAMP;
   #oSTW1.Bit_06_SETPOINT := #Temp_Eins AND #Temp_SEND.STW1.Bit_06_SETPOINT;
   #oSTW1.Bit_07_RESET := #Temp_Eins AND #Temp_SEND.STW1.Bit_07_RESET;
END_REGION

REGION Network 19: aktuelle Geschwindigkeit / CURR SPEED
   // ################################## oCURR_SPEED #################################
END_REGION

REGION Network 20 (STL): aktuelle Geschwindigkeit / CURR SPEED
   // PZD 2 - Drehzahlistwert
         L     #Temp_REC.SPEED;
         ITD;
         DTR;
         L     100.0;  // 16383= 4000HEX = 100%
         *R;
         L     16384.0;
         /R;
         L     100.0;  // nur 2-Nachkommastellen darstellen
         *R;
         TRUNC;
         ITD;
         DTR;
         L     100.0;
         /R;
         L     #Temp_Factor;
         /R;
         RND;
         T     #oCUR_SPEED;  // Istwert in m/min
END_REGION

REGION Network 21: Ausgänge PAW / OUTPUTS PAW
   // ##################################### PAW ######################################
END_REGION

REGION Network 22: OUT: G120 D Steuerwort 1 / Controlword 1 PAW
END_REGION

REGION Network 23: OUT: G120 D Soll-Drehzahl / Setpoint-Speed of rotation PAW
   RUNG wire#powerrail
      Move(in := #Temp_SEND.SPEED, out1 => #oPAW_SPEED)
   END_RUNG
   // the same network as SCL:
   #oPAW_SPEED := #Temp_SEND.SPEED;
END_REGION

REGION Network 24: STÖRUNGEN / FAULTS
   // ################################# STÖRUNGEN ########################## / #################################### FAULT ####################################
END_REGION

REGION Network 25: Störungen quittieren / reset Errors